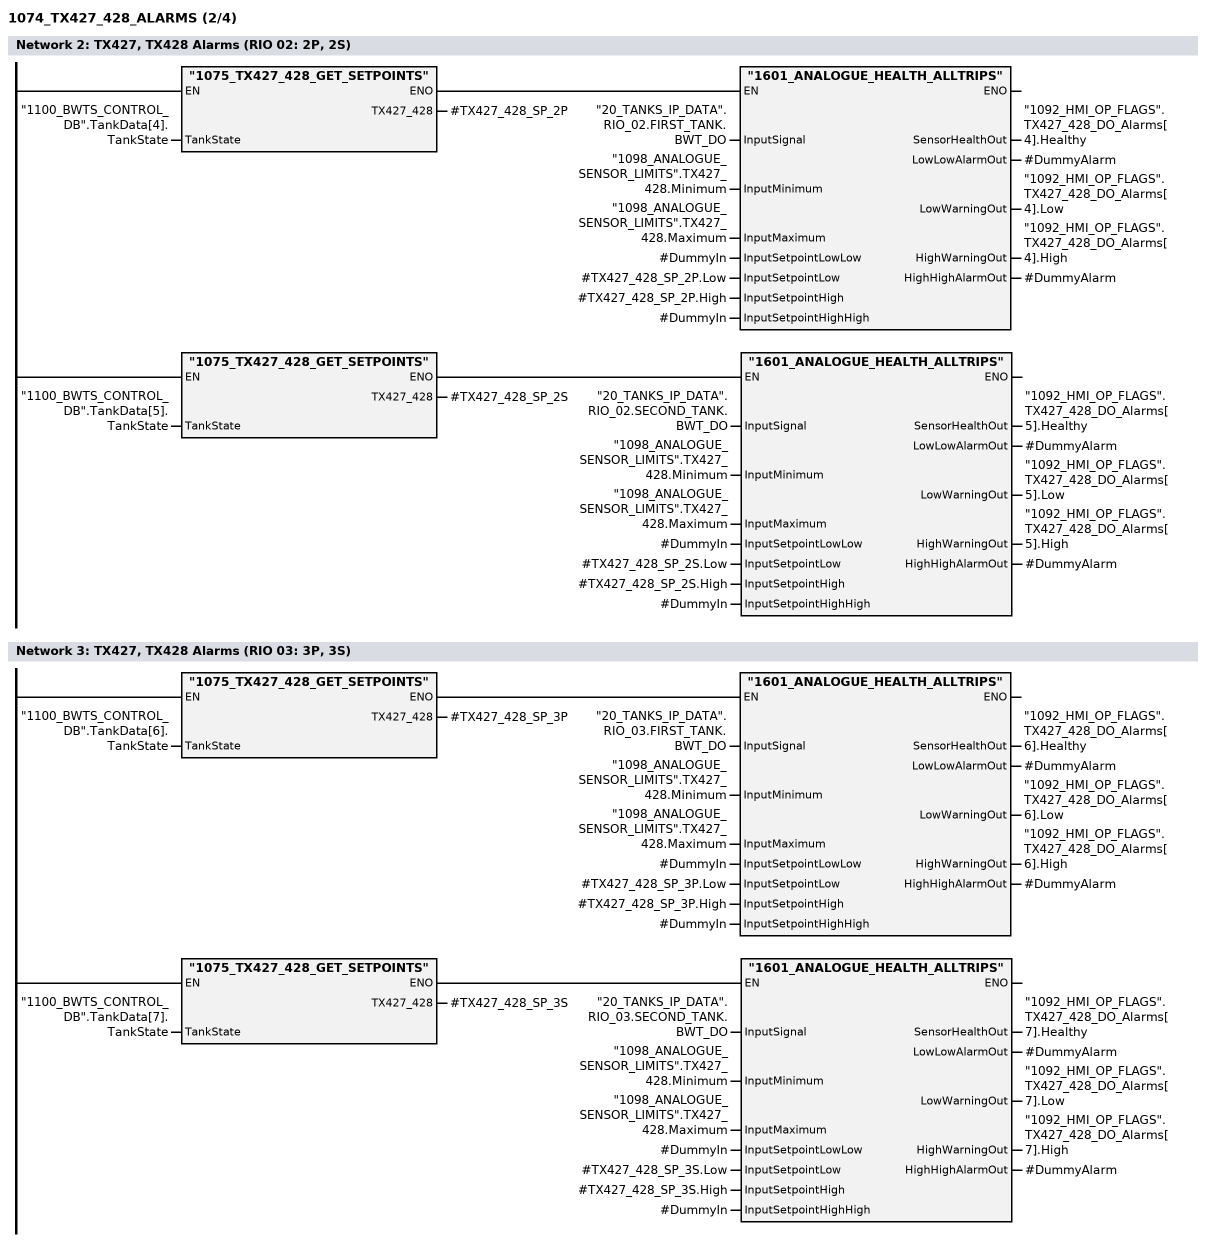
   RUNG wire#powerrail
      "1075_TX427_428_GET_SETPOINTS"(TankState := "1100_BWTS_CONTROL_DB".TankData[4].TankState, TX427_428 => #TX427_428_SP_2P)
      "1601_ANALOGUE_HEALTH_ALLTRIPS"(InputSignal := "20_TANKS_IP_DATA".RIO_02.FIRST_TANK.BWT_DO, InputMinimum := "1098_ANALOGUE_SENSOR_LIMITS".TX427_428.Minimum, InputMaximum := "1098_ANALOGUE_SENSOR_LIMITS".TX427_428.Maximum, InputSetpointLowLow := #DummyIn, InputSetpointLow := #TX427_428_SP_2P.Low, InputSetpointHigh := #TX427_428_SP_2P.High, InputSetpointHighHigh := #DummyIn, SensorHealthOut => "1092_HMI_OP_FLAGS".TX427_428_DO_Alarms[4].Healthy, LowLowAlarmOut => #DummyAlarm, LowWarningOut => "1092_HMI_OP_FLAGS".TX427_428_DO_Alarms[4].Low, HighWarningOut => "1092_HMI_OP_FLAGS".TX427_428_DO_Alarms[4].High, HighHighAlarmOut => #DummyAlarm)
   END_RUNG
   RUNG wire#powerrail
      "1075_TX427_428_GET_SETPOINTS"(TankState := "1100_BWTS_CONTROL_DB".TankData[5].TankState, TX427_428 => #TX427_428_SP_2S)
      "1601_ANALOGUE_HEALTH_ALLTRIPS"(InputSignal := "20_TANKS_IP_DATA".RIO_02.SECOND_TANK.BWT_DO, InputMinimum := "1098_ANALOGUE_SENSOR_LIMITS".TX427_428.Minimum, InputMaximum := "1098_ANALOGUE_SENSOR_LIMITS".TX427_428.Maximum, InputSetpointLowLow := #DummyIn, InputSetpointLow := #TX427_428_SP_2S.Low, InputSetpointHigh := #TX427_428_SP_2S.High, InputSetpointHighHigh := #DummyIn, SensorHealthOut => "1092_HMI_OP_FLAGS".TX427_428_DO_Alarms[5].Healthy, LowLowAlarmOut => #DummyAlarm, LowWarningOut => "1092_HMI_OP_FLAGS".TX427_428_DO_Alarms[5].Low, HighWarningOut => "1092_HMI_OP_FLAGS".TX427_428_DO_Alarms[5].High, HighHighAlarmOut => #DummyAlarm)
   END_RUNG
   // the same network as SCL:
   "1075_TX427_428_GET_SETPOINTS"(TankState := "1100_BWTS_CONTROL_DB".TankData[4].TankState,
                           TX427_428 => #TX427_428_SP_2P,
                           ENO => #_w1);
   IF #_w1 THEN
       "1601_ANALOGUE_HEALTH_ALLTRIPS"(InputSignal := "20_TANKS_IP_DATA".RIO_02.FIRST_TANK.BWT_DO,
                               InputMinimum := "1098_ANALOGUE_SENSOR_LIMITS".TX427_428.Minimum,
                               InputMaximum := "1098_ANALOGUE_SENSOR_LIMITS".TX427_428.Maximum,
                               InputSetpointLowLow := #DummyIn,
                               InputSetpointLow := #TX427_428_SP_2P.Low,
                               InputSetpointHigh := #TX427_428_SP_2P.High,
                               InputSetpointHighHigh := #DummyIn,
                               SensorHealthOut => "1092_HMI_OP_FLAGS".TX427_428_DO_Alarms[4].Healthy,
                               LowLowAlarmOut => #DummyAlarm,
                               LowWarningOut => "1092_HMI_OP_FLAGS".TX427_428_DO_Alarms[4].Low,
                               HighWarningOut => "1092_HMI_OP_FLAGS".TX427_428_DO_Alarms[4].High,
                               HighHighAlarmOut => #DummyAlarm);
   END_IF;
   "1075_TX427_428_GET_SETPOINTS"(TankState := "1100_BWTS_CONTROL_DB".TankData[5].TankState,
                           TX427_428 => #TX427_428_SP_2S,
                           ENO => #_w2);
   IF #_w2 THEN
       "1601_ANALOGUE_HEALTH_ALLTRIPS"(InputSignal := "20_TANKS_IP_DATA".RIO_02.SECOND_TANK.BWT_DO,
                               InputMinimum := "1098_ANALOGUE_SENSOR_LIMITS".TX427_428.Minimum,
                               InputMaximum := "1098_ANALOGUE_SENSOR_LIMITS".TX427_428.Maximum,
                               InputSetpointLowLow := #DummyIn,
                               InputSetpointLow := #TX427_428_SP_2S.Low,
                               InputSetpointHigh := #TX427_428_SP_2S.High,
                               InputSetpointHighHigh := #DummyIn,
                               SensorHealthOut => "1092_HMI_OP_FLAGS".TX427_428_DO_Alarms[5].Healthy,
                               LowLowAlarmOut => #DummyAlarm,
                               LowWarningOut => "1092_HMI_OP_FLAGS".TX427_428_DO_Alarms[5].Low,
                               HighWarningOut => "1092_HMI_OP_FLAGS".TX427_428_DO_Alarms[5].High,
                               HighHighAlarmOut => #DummyAlarm);
   END_IF;
END_REGION

REGION Network 3: TX427, TX428 Alarms (RIO 03: 3P, 3S)
   RUNG wire#powerrail
      "1075_TX427_428_GET_SETPOINTS"(TankState := "1100_BWTS_CONTROL_DB".TankData[6].TankState, TX427_428 => #TX427_428_SP_3P)
      "1601_ANALOGUE_HEALTH_ALLTRIPS"(InputSignal := "20_TANKS_IP_DATA".RIO_03.FIRST_TANK.BWT_DO, InputMinimum := "1098_ANALOGUE_SENSOR_LIMITS".TX427_428.Minimum, InputMaximum := "1098_ANALOGUE_SENSOR_LIMITS".TX427_428.Maximum, InputSetpointLowLow := #DummyIn, InputSetpointLow := #TX427_428_SP_3P.Low, InputSetpointHigh := #TX427_428_SP_3P.High, InputSetpointHighHigh := #DummyIn, SensorHealthOut => "1092_HMI_OP_FLAGS".TX427_428_DO_Alarms[6].Healthy, LowLowAlarmOut => #DummyAlarm, LowWarningOut => "1092_HMI_OP_FLAGS".TX427_428_DO_Alarms[6].Low, HighWarningOut => "1092_HMI_OP_FLAGS".TX427_428_DO_Alarms[6].High, HighHighAlarmOut => #DummyAlarm)
   END_RUNG
   RUNG wire#powerrail
      "1075_TX427_428_GET_SETPOINTS"(TankState := "1100_BWTS_CONTROL_DB".TankData[7].TankState, TX427_428 => #TX427_428_SP_3S)
      "1601_ANALOGUE_HEALTH_ALLTRIPS"(InputSignal := "20_TANKS_IP_DATA".RIO_03.SECOND_TANK.BWT_DO, InputMinimum := "1098_ANALOGUE_SENSOR_LIMITS".TX427_428.Minimum, InputMaximum := "1098_ANALOGUE_SENSOR_LIMITS".TX427_428.Maximum, InputSetpointLowLow := #DummyIn, InputSetpointLow := #TX427_428_SP_3S.Low, InputSetpointHigh := #TX427_428_SP_3S.High, InputSetpointHighHigh := #DummyIn, SensorHealthOut => "1092_HMI_OP_FLAGS".TX427_428_DO_Alarms[7].Healthy, LowLowAlarmOut => #DummyAlarm, LowWarningOut => "1092_HMI_OP_FLAGS".TX427_428_DO_Alarms[7].Low, HighWarningOut => "1092_HMI_OP_FLAGS".TX427_428_DO_Alarms[7].High, HighHighAlarmOut => #DummyAlarm)
   END_RUNG
   // the same network as SCL:
   "1075_TX427_428_GET_SETPOINTS"(TankState := "1100_BWTS_CONTROL_DB".TankData[6].TankState,
                           TX427_428 => #TX427_428_SP_3P,
                           ENO => #_w1);
   IF #_w1 THEN
       "1601_ANALOGUE_HEALTH_ALLTRIPS"(InputSignal := "20_TANKS_IP_DATA".RIO_03.FIRST_TANK.BWT_DO,
                               InputMinimum := "1098_ANALOGUE_SENSOR_LIMITS".TX427_428.Minimum,
                               InputMaximum := "1098_ANALOGUE_SENSOR_LIMITS".TX427_428.Maximum,
                               InputSetpointLowLow := #DummyIn,
                               InputSetpointLow := #TX427_428_SP_3P.Low,
                               InputSetpointHigh := #TX427_428_SP_3P.High,
                               InputSetpointHighHigh := #DummyIn,
                               SensorHealthOut => "1092_HMI_OP_FLAGS".TX427_428_DO_Alarms[6].Healthy,
                               LowLowAlarmOut => #DummyAlarm,
                               LowWarningOut => "1092_HMI_OP_FLAGS".TX427_428_DO_Alarms[6].Low,
                               HighWarningOut => "1092_HMI_OP_FLAGS".TX427_428_DO_Alarms[6].High,
                               HighHighAlarmOut => #DummyAlarm);
   END_IF;
   "1075_TX427_428_GET_SETPOINTS"(TankState := "1100_BWTS_CONTROL_DB".TankData[7].TankState,
                           TX427_428 => #TX427_428_SP_3S,
                           ENO => #_w2);
   IF #_w2 THEN
       "1601_ANALOGUE_HEALTH_ALLTRIPS"(InputSignal := "20_TANKS_IP_DATA".RIO_03.SECOND_TANK.BWT_DO,
                               InputMinimum := "1098_ANALOGUE_SENSOR_LIMITS".TX427_428.Minimum,
                               InputMaximum := "1098_ANALOGUE_SENSOR_LIMITS".TX427_428.Maximum,
                               InputSetpointLowLow := #DummyIn,
                               InputSetpointLow := #TX427_428_SP_3S.Low,
                               InputSetpointHigh := #TX427_428_SP_3S.High,
                               InputSetpointHighHigh := #DummyIn,
                               SensorHealthOut => "1092_HMI_OP_FLAGS".TX427_428_DO_Alarms[7].Healthy,
                               LowLowAlarmOut => #DummyAlarm,
                               LowWarningOut => "1092_HMI_OP_FLAGS".TX427_428_DO_Alarms[7].Low,
                               HighWarningOut => "1092_HMI_OP_FLAGS".TX427_428_DO_Alarms[7].High,
                               HighHighAlarmOut => #DummyAlarm);
   END_IF;
END_REGION

REGION Network 4: TX427, TX428 Alarms (RIO 04: 4P, 4S)
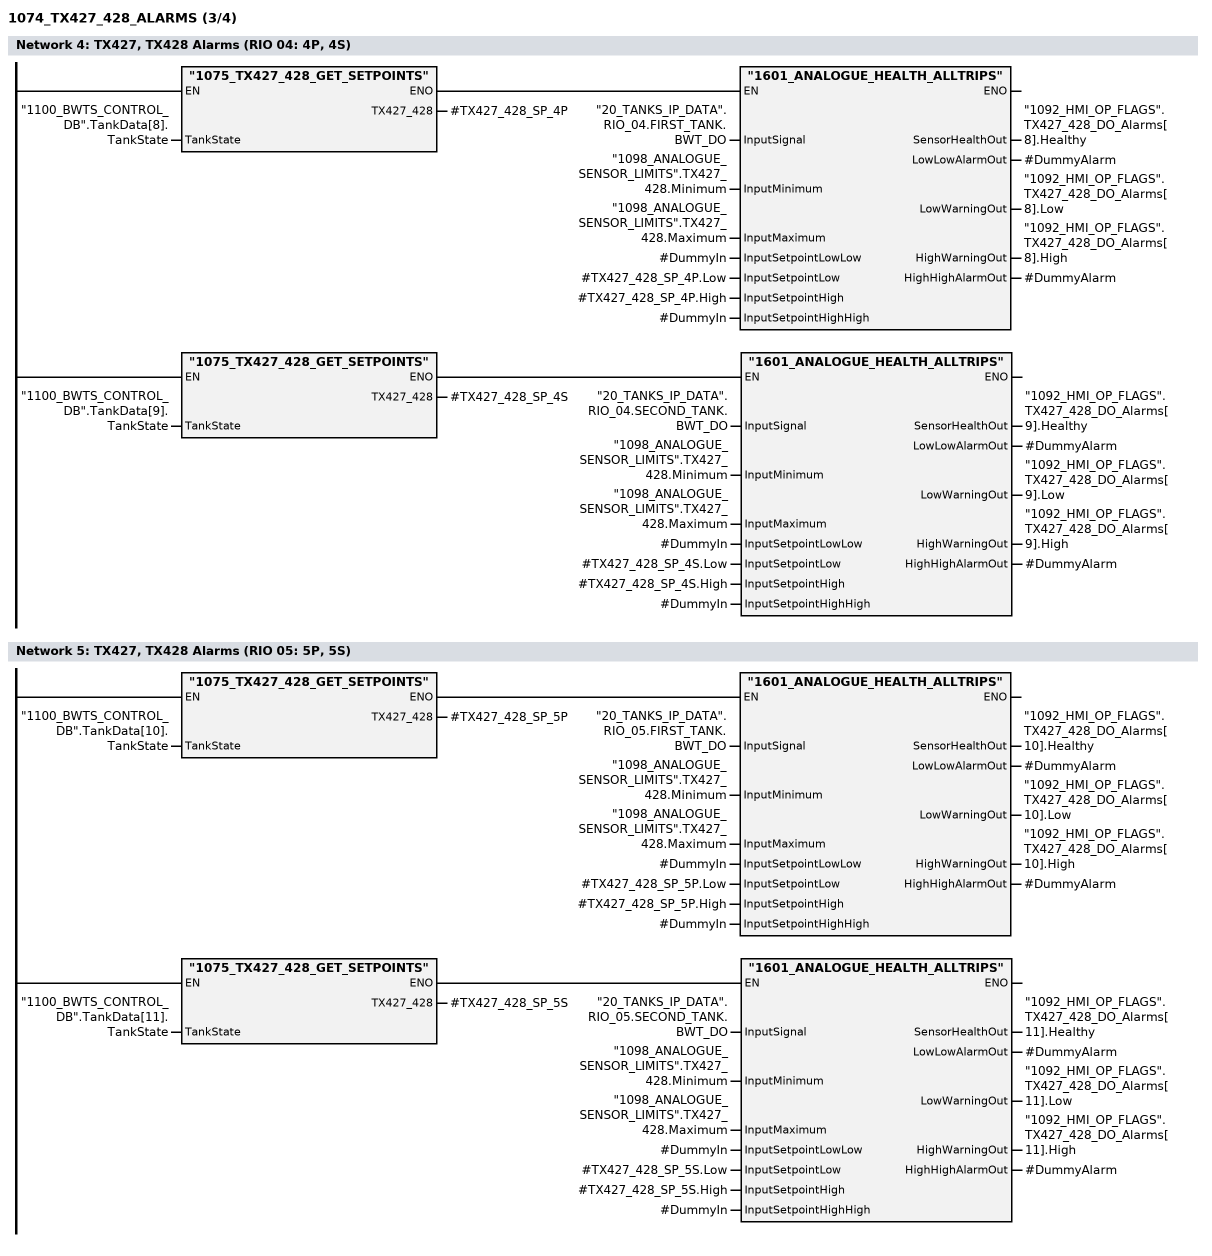
   RUNG wire#powerrail
      "1075_TX427_428_GET_SETPOINTS"(TankState := "1100_BWTS_CONTROL_DB".TankData[8].TankState, TX427_428 => #TX427_428_SP_4P)
      "1601_ANALOGUE_HEALTH_ALLTRIPS"(InputSignal := "20_TANKS_IP_DATA".RIO_04.FIRST_TANK.BWT_DO, InputMinimum := "1098_ANALOGUE_SENSOR_LIMITS".TX427_428.Minimum, InputMaximum := "1098_ANALOGUE_SENSOR_LIMITS".TX427_428.Maximum, InputSetpointLowLow := #DummyIn, InputSetpointLow := #TX427_428_SP_4P.Low, InputSetpointHigh := #TX427_428_SP_4P.High, InputSetpointHighHigh := #DummyIn, SensorHealthOut => "1092_HMI_OP_FLAGS".TX427_428_DO_Alarms[8].Healthy, LowLowAlarmOut => #DummyAlarm, LowWarningOut => "1092_HMI_OP_FLAGS".TX427_428_DO_Alarms[8].Low, HighWarningOut => "1092_HMI_OP_FLAGS".TX427_428_DO_Alarms[8].High, HighHighAlarmOut => #DummyAlarm)
   END_RUNG
   RUNG wire#powerrail
      "1075_TX427_428_GET_SETPOINTS"(TankState := "1100_BWTS_CONTROL_DB".TankData[9].TankState, TX427_428 => #TX427_428_SP_4S)
      "1601_ANALOGUE_HEALTH_ALLTRIPS"(InputSignal := "20_TANKS_IP_DATA".RIO_04.SECOND_TANK.BWT_DO, InputMinimum := "1098_ANALOGUE_SENSOR_LIMITS".TX427_428.Minimum, InputMaximum := "1098_ANALOGUE_SENSOR_LIMITS".TX427_428.Maximum, InputSetpointLowLow := #DummyIn, InputSetpointLow := #TX427_428_SP_4S.Low, InputSetpointHigh := #TX427_428_SP_4S.High, InputSetpointHighHigh := #DummyIn, SensorHealthOut => "1092_HMI_OP_FLAGS".TX427_428_DO_Alarms[9].Healthy, LowLowAlarmOut => #DummyAlarm, LowWarningOut => "1092_HMI_OP_FLAGS".TX427_428_DO_Alarms[9].Low, HighWarningOut => "1092_HMI_OP_FLAGS".TX427_428_DO_Alarms[9].High, HighHighAlarmOut => #DummyAlarm)
   END_RUNG
   // the same network as SCL:
   "1075_TX427_428_GET_SETPOINTS"(TankState := "1100_BWTS_CONTROL_DB".TankData[8].TankState,
                           TX427_428 => #TX427_428_SP_4P,
                           ENO => #_w1);
   IF #_w1 THEN
       "1601_ANALOGUE_HEALTH_ALLTRIPS"(InputSignal := "20_TANKS_IP_DATA".RIO_04.FIRST_TANK.BWT_DO,
                               InputMinimum := "1098_ANALOGUE_SENSOR_LIMITS".TX427_428.Minimum,
                               InputMaximum := "1098_ANALOGUE_SENSOR_LIMITS".TX427_428.Maximum,
                               InputSetpointLowLow := #DummyIn,
                               InputSetpointLow := #TX427_428_SP_4P.Low,
                               InputSetpointHigh := #TX427_428_SP_4P.High,
                               InputSetpointHighHigh := #DummyIn,
                               SensorHealthOut => "1092_HMI_OP_FLAGS".TX427_428_DO_Alarms[8].Healthy,
                               LowLowAlarmOut => #DummyAlarm,
                               LowWarningOut => "1092_HMI_OP_FLAGS".TX427_428_DO_Alarms[8].Low,
                               HighWarningOut => "1092_HMI_OP_FLAGS".TX427_428_DO_Alarms[8].High,
                               HighHighAlarmOut => #DummyAlarm);
   END_IF;
   "1075_TX427_428_GET_SETPOINTS"(TankState := "1100_BWTS_CONTROL_DB".TankData[9].TankState,
                           TX427_428 => #TX427_428_SP_4S,
                           ENO => #_w2);
   IF #_w2 THEN
       "1601_ANALOGUE_HEALTH_ALLTRIPS"(InputSignal := "20_TANKS_IP_DATA".RIO_04.SECOND_TANK.BWT_DO,
                               InputMinimum := "1098_ANALOGUE_SENSOR_LIMITS".TX427_428.Minimum,
                               InputMaximum := "1098_ANALOGUE_SENSOR_LIMITS".TX427_428.Maximum,
                               InputSetpointLowLow := #DummyIn,
                               InputSetpointLow := #TX427_428_SP_4S.Low,
                               InputSetpointHigh := #TX427_428_SP_4S.High,
                               InputSetpointHighHigh := #DummyIn,
                               SensorHealthOut => "1092_HMI_OP_FLAGS".TX427_428_DO_Alarms[9].Healthy,
                               LowLowAlarmOut => #DummyAlarm,
                               LowWarningOut => "1092_HMI_OP_FLAGS".TX427_428_DO_Alarms[9].Low,
                               HighWarningOut => "1092_HMI_OP_FLAGS".TX427_428_DO_Alarms[9].High,
                               HighHighAlarmOut => #DummyAlarm);
   END_IF;
END_REGION

REGION Network 5: TX427, TX428 Alarms (RIO 05: 5P, 5S)
   RUNG wire#powerrail
      "1075_TX427_428_GET_SETPOINTS"(TankState := "1100_BWTS_CONTROL_DB".TankData[10].TankState, TX427_428 => #TX427_428_SP_5P)
      "1601_ANALOGUE_HEALTH_ALLTRIPS"(InputSignal := "20_TANKS_IP_DATA".RIO_05.FIRST_TANK.BWT_DO, InputMinimum := "1098_ANALOGUE_SENSOR_LIMITS".TX427_428.Minimum, InputMaximum := "1098_ANALOGUE_SENSOR_LIMITS".TX427_428.Maximum, InputSetpointLowLow := #DummyIn, InputSetpointLow := #TX427_428_SP_5P.Low, InputSetpointHigh := #TX427_428_SP_5P.High, InputSetpointHighHigh := #DummyIn, SensorHealthOut => "1092_HMI_OP_FLAGS".TX427_428_DO_Alarms[10].Healthy, LowLowAlarmOut => #DummyAlarm, LowWarningOut => "1092_HMI_OP_FLAGS".TX427_428_DO_Alarms[10].Low, HighWarningOut => "1092_HMI_OP_FLAGS".TX427_428_DO_Alarms[10].High, HighHighAlarmOut => #DummyAlarm)
   END_RUNG
   RUNG wire#powerrail
      "1075_TX427_428_GET_SETPOINTS"(TankState := "1100_BWTS_CONTROL_DB".TankData[11].TankState, TX427_428 => #TX427_428_SP_5S)
      "1601_ANALOGUE_HEALTH_ALLTRIPS"(InputSignal := "20_TANKS_IP_DATA".RIO_05.SECOND_TANK.BWT_DO, InputMinimum := "1098_ANALOGUE_SENSOR_LIMITS".TX427_428.Minimum, InputMaximum := "1098_ANALOGUE_SENSOR_LIMITS".TX427_428.Maximum, InputSetpointLowLow := #DummyIn, InputSetpointLow := #TX427_428_SP_5S.Low, InputSetpointHigh := #TX427_428_SP_5S.High, InputSetpointHighHigh := #DummyIn, SensorHealthOut => "1092_HMI_OP_FLAGS".TX427_428_DO_Alarms[11].Healthy, LowLowAlarmOut => #DummyAlarm, LowWarningOut => "1092_HMI_OP_FLAGS".TX427_428_DO_Alarms[11].Low, HighWarningOut => "1092_HMI_OP_FLAGS".TX427_428_DO_Alarms[11].High, HighHighAlarmOut => #DummyAlarm)
   END_RUNG
   // the same network as SCL:
   "1075_TX427_428_GET_SETPOINTS"(TankState := "1100_BWTS_CONTROL_DB".TankData[10].TankState,
                           TX427_428 => #TX427_428_SP_5P,
                           ENO => #_w1);
   IF #_w1 THEN
       "1601_ANALOGUE_HEALTH_ALLTRIPS"(InputSignal := "20_TANKS_IP_DATA".RIO_05.FIRST_TANK.BWT_DO,
                               InputMinimum := "1098_ANALOGUE_SENSOR_LIMITS".TX427_428.Minimum,
                               InputMaximum := "1098_ANALOGUE_SENSOR_LIMITS".TX427_428.Maximum,
                               InputSetpointLowLow := #DummyIn,
                               InputSetpointLow := #TX427_428_SP_5P.Low,
                               InputSetpointHigh := #TX427_428_SP_5P.High,
                               InputSetpointHighHigh := #DummyIn,
                               SensorHealthOut => "1092_HMI_OP_FLAGS".TX427_428_DO_Alarms[10].Healthy,
                               LowLowAlarmOut => #DummyAlarm,
                               LowWarningOut => "1092_HMI_OP_FLAGS".TX427_428_DO_Alarms[10].Low,
                               HighWarningOut => "1092_HMI_OP_FLAGS".TX427_428_DO_Alarms[10].High,
                               HighHighAlarmOut => #DummyAlarm);
   END_IF;
   "1075_TX427_428_GET_SETPOINTS"(TankState := "1100_BWTS_CONTROL_DB".TankData[11].TankState,
                           TX427_428 => #TX427_428_SP_5S,
                           ENO => #_w2);
   IF #_w2 THEN
       "1601_ANALOGUE_HEALTH_ALLTRIPS"(InputSignal := "20_TANKS_IP_DATA".RIO_05.SECOND_TANK.BWT_DO,
                               InputMinimum := "1098_ANALOGUE_SENSOR_LIMITS".TX427_428.Minimum,
                               InputMaximum := "1098_ANALOGUE_SENSOR_LIMITS".TX427_428.Maximum,
                               InputSetpointLowLow := #DummyIn,
                               InputSetpointLow := #TX427_428_SP_5S.Low,
                               InputSetpointHigh := #TX427_428_SP_5S.High,
                               InputSetpointHighHigh := #DummyIn,
                               SensorHealthOut => "1092_HMI_OP_FLAGS".TX427_428_DO_Alarms[11].Healthy,
                               LowLowAlarmOut => #DummyAlarm,
                               LowWarningOut => "1092_HMI_OP_FLAGS".TX427_428_DO_Alarms[11].Low,
                               HighWarningOut => "1092_HMI_OP_FLAGS".TX427_428_DO_Alarms[11].High,
                               HighHighAlarmOut => #DummyAlarm);
   END_IF;
END_REGION

REGION Network 6: TX427, TX428 Alarms (RIO 06: 6P, 6S)
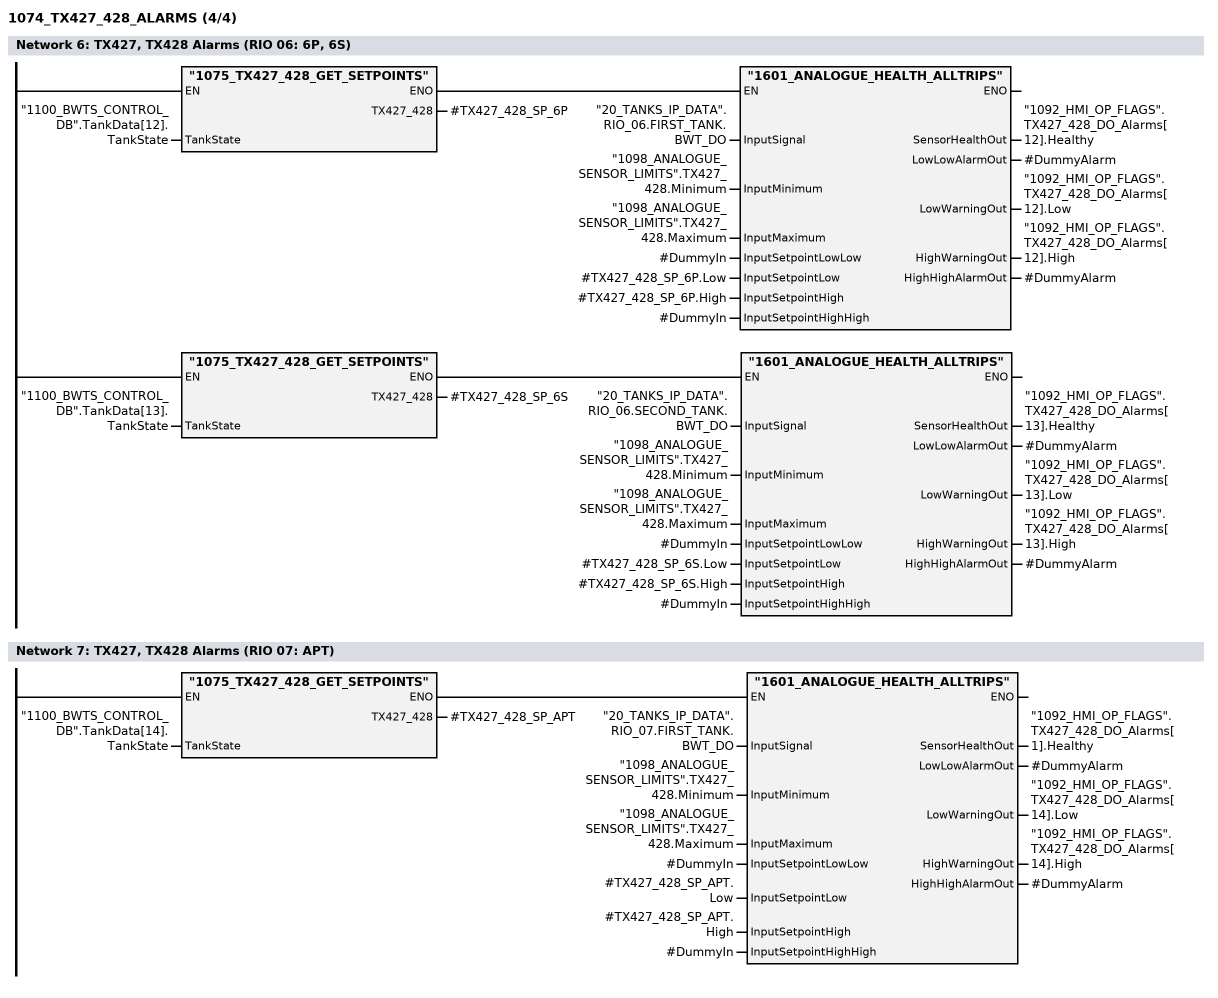
   RUNG wire#powerrail
      "1075_TX427_428_GET_SETPOINTS"(TankState := "1100_BWTS_CONTROL_DB".TankData[12].TankState, TX427_428 => #TX427_428_SP_6P)
      "1601_ANALOGUE_HEALTH_ALLTRIPS"(InputSignal := "20_TANKS_IP_DATA".RIO_06.FIRST_TANK.BWT_DO, InputMinimum := "1098_ANALOGUE_SENSOR_LIMITS".TX427_428.Minimum, InputMaximum := "1098_ANALOGUE_SENSOR_LIMITS".TX427_428.Maximum, InputSetpointLowLow := #DummyIn, InputSetpointLow := #TX427_428_SP_6P.Low, InputSetpointHigh := #TX427_428_SP_6P.High, InputSetpointHighHigh := #DummyIn, SensorHealthOut => "1092_HMI_OP_FLAGS".TX427_428_DO_Alarms[12].Healthy, LowLowAlarmOut => #DummyAlarm, LowWarningOut => "1092_HMI_OP_FLAGS".TX427_428_DO_Alarms[12].Low, HighWarningOut => "1092_HMI_OP_FLAGS".TX427_428_DO_Alarms[12].High, HighHighAlarmOut => #DummyAlarm)
   END_RUNG
   RUNG wire#powerrail
      "1075_TX427_428_GET_SETPOINTS"(TankState := "1100_BWTS_CONTROL_DB".TankData[13].TankState, TX427_428 => #TX427_428_SP_6S)
      "1601_ANALOGUE_HEALTH_ALLTRIPS"(InputSignal := "20_TANKS_IP_DATA".RIO_06.SECOND_TANK.BWT_DO, InputMinimum := "1098_ANALOGUE_SENSOR_LIMITS".TX427_428.Minimum, InputMaximum := "1098_ANALOGUE_SENSOR_LIMITS".TX427_428.Maximum, InputSetpointLowLow := #DummyIn, InputSetpointLow := #TX427_428_SP_6S.Low, InputSetpointHigh := #TX427_428_SP_6S.High, InputSetpointHighHigh := #DummyIn, SensorHealthOut => "1092_HMI_OP_FLAGS".TX427_428_DO_Alarms[13].Healthy, LowLowAlarmOut => #DummyAlarm, LowWarningOut => "1092_HMI_OP_FLAGS".TX427_428_DO_Alarms[13].Low, HighWarningOut => "1092_HMI_OP_FLAGS".TX427_428_DO_Alarms[13].High, HighHighAlarmOut => #DummyAlarm)
   END_RUNG
   // the same network as SCL:
   "1075_TX427_428_GET_SETPOINTS"(TankState := "1100_BWTS_CONTROL_DB".TankData[12].TankState,
                           TX427_428 => #TX427_428_SP_6P,
                           ENO => #_w1);
   IF #_w1 THEN
       "1601_ANALOGUE_HEALTH_ALLTRIPS"(InputSignal := "20_TANKS_IP_DATA".RIO_06.FIRST_TANK.BWT_DO,
                               InputMinimum := "1098_ANALOGUE_SENSOR_LIMITS".TX427_428.Minimum,
                               InputMaximum := "1098_ANALOGUE_SENSOR_LIMITS".TX427_428.Maximum,
                               InputSetpointLowLow := #DummyIn,
                               InputSetpointLow := #TX427_428_SP_6P.Low,
                               InputSetpointHigh := #TX427_428_SP_6P.High,
                               InputSetpointHighHigh := #DummyIn,
                               SensorHealthOut => "1092_HMI_OP_FLAGS".TX427_428_DO_Alarms[12].Healthy,
                               LowLowAlarmOut => #DummyAlarm,
                               LowWarningOut => "1092_HMI_OP_FLAGS".TX427_428_DO_Alarms[12].Low,
                               HighWarningOut => "1092_HMI_OP_FLAGS".TX427_428_DO_Alarms[12].High,
                               HighHighAlarmOut => #DummyAlarm);
   END_IF;
   "1075_TX427_428_GET_SETPOINTS"(TankState := "1100_BWTS_CONTROL_DB".TankData[13].TankState,
                           TX427_428 => #TX427_428_SP_6S,
                           ENO => #_w2);
   IF #_w2 THEN
       "1601_ANALOGUE_HEALTH_ALLTRIPS"(InputSignal := "20_TANKS_IP_DATA".RIO_06.SECOND_TANK.BWT_DO,
                               InputMinimum := "1098_ANALOGUE_SENSOR_LIMITS".TX427_428.Minimum,
                               InputMaximum := "1098_ANALOGUE_SENSOR_LIMITS".TX427_428.Maximum,
                               InputSetpointLowLow := #DummyIn,
                               InputSetpointLow := #TX427_428_SP_6S.Low,
                               InputSetpointHigh := #TX427_428_SP_6S.High,
                               InputSetpointHighHigh := #DummyIn,
                               SensorHealthOut => "1092_HMI_OP_FLAGS".TX427_428_DO_Alarms[13].Healthy,
                               LowLowAlarmOut => #DummyAlarm,
                               LowWarningOut => "1092_HMI_OP_FLAGS".TX427_428_DO_Alarms[13].Low,
                               HighWarningOut => "1092_HMI_OP_FLAGS".TX427_428_DO_Alarms[13].High,
                               HighHighAlarmOut => #DummyAlarm);
   END_IF;
END_REGION

REGION Network 7: TX427, TX428 Alarms (RIO 07: APT)
   RUNG wire#powerrail
      "1075_TX427_428_GET_SETPOINTS"(TankState := "1100_BWTS_CONTROL_DB".TankData[14].TankState, TX427_428 => #TX427_428_SP_APT)
      "1601_ANALOGUE_HEALTH_ALLTRIPS"(InputSignal := "20_TANKS_IP_DATA".RIO_07.FIRST_TANK.BWT_DO, InputMinimum := "1098_ANALOGUE_SENSOR_LIMITS".TX427_428.Minimum, InputMaximum := "1098_ANALOGUE_SENSOR_LIMITS".TX427_428.Maximum, InputSetpointLowLow := #DummyIn, InputSetpointLow := #TX427_428_SP_APT.Low, InputSetpointHigh := #TX427_428_SP_APT.High, InputSetpointHighHigh := #DummyIn, SensorHealthOut => "1092_HMI_OP_FLAGS".TX427_428_DO_Alarms[1].Healthy, LowLowAlarmOut => #DummyAlarm, LowWarningOut => "1092_HMI_OP_FLAGS".TX427_428_DO_Alarms[14].Low, HighWarningOut => "1092_HMI_OP_FLAGS".TX427_428_DO_Alarms[14].High, HighHighAlarmOut => #DummyAlarm)
   END_RUNG
   // the same network as SCL:
   "1075_TX427_428_GET_SETPOINTS"(TankState := "1100_BWTS_CONTROL_DB".TankData[14].TankState,
                           TX427_428 => #TX427_428_SP_APT,
                           ENO => #_w1);
   IF #_w1 THEN
       "1601_ANALOGUE_HEALTH_ALLTRIPS"(InputSignal := "20_TANKS_IP_DATA".RIO_07.FIRST_TANK.BWT_DO,
                               InputMinimum := "1098_ANALOGUE_SENSOR_LIMITS".TX427_428.Minimum,
                               InputMaximum := "1098_ANALOGUE_SENSOR_LIMITS".TX427_428.Maximum,
                               InputSetpointLowLow := #DummyIn,
                               InputSetpointLow := #TX427_428_SP_APT.Low,
                               InputSetpointHigh := #TX427_428_SP_APT.High,
                               InputSetpointHighHigh := #DummyIn,
                               SensorHealthOut => "1092_HMI_OP_FLAGS".TX427_428_DO_Alarms[1].Healthy,
                               LowLowAlarmOut => #DummyAlarm,
                               LowWarningOut => "1092_HMI_OP_FLAGS".TX427_428_DO_Alarms[14].Low,
                               HighWarningOut => "1092_HMI_OP_FLAGS".TX427_428_DO_Alarms[14].High,
                               HighHighAlarmOut => #DummyAlarm);
   END_IF;
END_REGION
END_FUNCTION

FUNCTION "1075_TX427_428_GET_SETPOINTS" : Void   // FC1075, SCL
{ S7_Optimized_Access := 'TRUE' }
VERSION : 0.1
   VAR_INPUT
      TankState : Int;
   END_VAR
   VAR_OUTPUT
      TX427_428 : "ANALOG_SENSOR_SETPOINTS";
   END_VAR
   VAR CONSTANT
      TankState_Init : Int := 1000;
      TankState_PreDwell : Int := 1001;
      TankState_DeOx : Int := 1002;
      TankState_MidDwell : Int := 1003;
      TankState_ReOx : Int := 1004;
      TankState_PostDwell : Int := 1005;
      TankState_Done : Int := 1006;
   END_VAR
BEGIN
   (* This function is required to define the setpoints of the DO sensors based on the current state.
       The alarms shall use differing setpoints in different phases defined as:
       DEOX alarm setpoints if in DeOx, or Mid-Dwell
       REOX alarm setpoints if in PreDwell, Reox, or PostDwell (All others values) *)

   IF #TankState = #TankState_DeOx OR #TankState = #TankState_MidDwell THEN
       #TX427_428 := "1094_ANALOGUE_SENSOR_SETPOINTS".TX427_428_DEOX;
   ELSE
       #TX427_428 := "1094_ANALOGUE_SENSOR_SETPOINTS".TX427_428_REOX;
   END_IF;
END_FUNCTION

FUNCTION "1076_LS425_442_ALARMS" : Void   // FC1076, LAD
{ S7_Optimized_Access := 'TRUE' }
VERSION : 0.1
// Alarm wrapper function for BWT Level Switch on each tank.
   VAR CONSTANT
      InputTripLevel : Bool;   // The input trip level for this function, if the input is equal to this digital value, trip the alarm.
   END_VAR
BEGIN

REGION Network 1: LS425, LS442 Alarms (RIO 01: FPT. 1P, 1S)
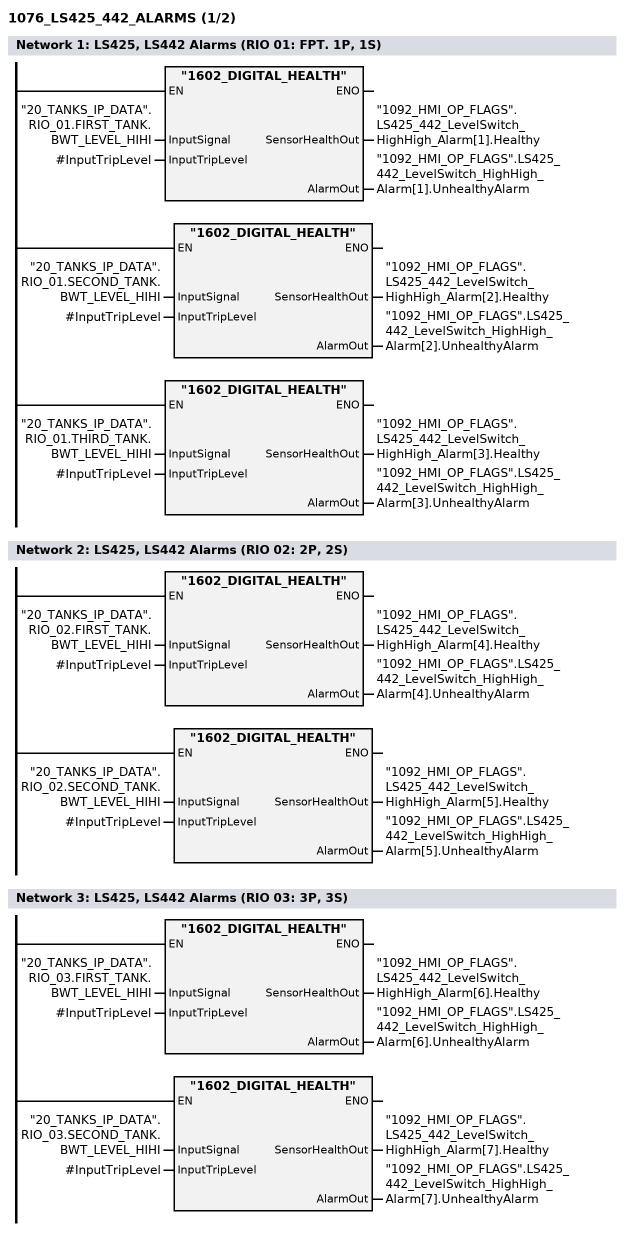
   RUNG wire#powerrail
      "1602_DIGITAL_HEALTH"(InputSignal := "20_TANKS_IP_DATA".RIO_01.FIRST_TANK.BWT_LEVEL_HIHI, InputTripLevel := #InputTripLevel, SensorHealthOut => "1092_HMI_OP_FLAGS".LS425_442_LevelSwitch_HighHigh_Alarm[1].Healthy, AlarmOut => "1092_HMI_OP_FLAGS".LS425_442_LevelSwitch_HighHigh_Alarm[1].UnhealthyAlarm)
   END_RUNG
   RUNG wire#powerrail
      "1602_DIGITAL_HEALTH"(InputSignal := "20_TANKS_IP_DATA".RIO_01.SECOND_TANK.BWT_LEVEL_HIHI, InputTripLevel := #InputTripLevel, SensorHealthOut => "1092_HMI_OP_FLAGS".LS425_442_LevelSwitch_HighHigh_Alarm[2].Healthy, AlarmOut => "1092_HMI_OP_FLAGS".LS425_442_LevelSwitch_HighHigh_Alarm[2].UnhealthyAlarm)
   END_RUNG
   RUNG wire#powerrail
      "1602_DIGITAL_HEALTH"(InputSignal := "20_TANKS_IP_DATA".RIO_01.THIRD_TANK.BWT_LEVEL_HIHI, InputTripLevel := #InputTripLevel, SensorHealthOut => "1092_HMI_OP_FLAGS".LS425_442_LevelSwitch_HighHigh_Alarm[3].Healthy, AlarmOut => "1092_HMI_OP_FLAGS".LS425_442_LevelSwitch_HighHigh_Alarm[3].UnhealthyAlarm)
   END_RUNG
   // the same network as SCL:
   "1602_DIGITAL_HEALTH"(InputSignal := "20_TANKS_IP_DATA".RIO_01.FIRST_TANK.BWT_LEVEL_HIHI,
                         InputTripLevel := #InputTripLevel,
                         SensorHealthOut => "1092_HMI_OP_FLAGS".LS425_442_LevelSwitch_HighHigh_Alarm[1].Healthy,
                         AlarmOut => "1092_HMI_OP_FLAGS".LS425_442_LevelSwitch_HighHigh_Alarm[1].UnhealthyAlarm);
   "1602_DIGITAL_HEALTH"(InputSignal := "20_TANKS_IP_DATA".RIO_01.SECOND_TANK.BWT_LEVEL_HIHI,
                         InputTripLevel := #InputTripLevel,
                         SensorHealthOut => "1092_HMI_OP_FLAGS".LS425_442_LevelSwitch_HighHigh_Alarm[2].Healthy,
                         AlarmOut => "1092_HMI_OP_FLAGS".LS425_442_LevelSwitch_HighHigh_Alarm[2].UnhealthyAlarm);
   "1602_DIGITAL_HEALTH"(InputSignal := "20_TANKS_IP_DATA".RIO_01.THIRD_TANK.BWT_LEVEL_HIHI,
                         InputTripLevel := #InputTripLevel,
                         SensorHealthOut => "1092_HMI_OP_FLAGS".LS425_442_LevelSwitch_HighHigh_Alarm[3].Healthy,
                         AlarmOut => "1092_HMI_OP_FLAGS".LS425_442_LevelSwitch_HighHigh_Alarm[3].UnhealthyAlarm);
END_REGION

REGION Network 2: LS425, LS442 Alarms (RIO 02: 2P, 2S)
   RUNG wire#powerrail
      "1602_DIGITAL_HEALTH"(InputSignal := "20_TANKS_IP_DATA".RIO_02.FIRST_TANK.BWT_LEVEL_HIHI, InputTripLevel := #InputTripLevel, SensorHealthOut => "1092_HMI_OP_FLAGS".LS425_442_LevelSwitch_HighHigh_Alarm[4].Healthy, AlarmOut => "1092_HMI_OP_FLAGS".LS425_442_LevelSwitch_HighHigh_Alarm[4].UnhealthyAlarm)
   END_RUNG
   RUNG wire#powerrail
      "1602_DIGITAL_HEALTH"(InputSignal := "20_TANKS_IP_DATA".RIO_02.SECOND_TANK.BWT_LEVEL_HIHI, InputTripLevel := #InputTripLevel, SensorHealthOut => "1092_HMI_OP_FLAGS".LS425_442_LevelSwitch_HighHigh_Alarm[5].Healthy, AlarmOut => "1092_HMI_OP_FLAGS".LS425_442_LevelSwitch_HighHigh_Alarm[5].UnhealthyAlarm)
   END_RUNG
   // the same network as SCL:
   "1602_DIGITAL_HEALTH"(InputSignal := "20_TANKS_IP_DATA".RIO_02.FIRST_TANK.BWT_LEVEL_HIHI,
                         InputTripLevel := #InputTripLevel,
                         SensorHealthOut => "1092_HMI_OP_FLAGS".LS425_442_LevelSwitch_HighHigh_Alarm[4].Healthy,
                         AlarmOut => "1092_HMI_OP_FLAGS".LS425_442_LevelSwitch_HighHigh_Alarm[4].UnhealthyAlarm);
   "1602_DIGITAL_HEALTH"(InputSignal := "20_TANKS_IP_DATA".RIO_02.SECOND_TANK.BWT_LEVEL_HIHI,
                         InputTripLevel := #InputTripLevel,
                         SensorHealthOut => "1092_HMI_OP_FLAGS".LS425_442_LevelSwitch_HighHigh_Alarm[5].Healthy,
                         AlarmOut => "1092_HMI_OP_FLAGS".LS425_442_LevelSwitch_HighHigh_Alarm[5].UnhealthyAlarm);
END_REGION

REGION Network 3: LS425, LS442 Alarms (RIO 03: 3P, 3S)
   RUNG wire#powerrail
      "1602_DIGITAL_HEALTH"(InputSignal := "20_TANKS_IP_DATA".RIO_03.FIRST_TANK.BWT_LEVEL_HIHI, InputTripLevel := #InputTripLevel, SensorHealthOut => "1092_HMI_OP_FLAGS".LS425_442_LevelSwitch_HighHigh_Alarm[6].Healthy, AlarmOut => "1092_HMI_OP_FLAGS".LS425_442_LevelSwitch_HighHigh_Alarm[6].UnhealthyAlarm)
   END_RUNG
   RUNG wire#powerrail
      "1602_DIGITAL_HEALTH"(InputSignal := "20_TANKS_IP_DATA".RIO_03.SECOND_TANK.BWT_LEVEL_HIHI, InputTripLevel := #InputTripLevel, SensorHealthOut => "1092_HMI_OP_FLAGS".LS425_442_LevelSwitch_HighHigh_Alarm[7].Healthy, AlarmOut => "1092_HMI_OP_FLAGS".LS425_442_LevelSwitch_HighHigh_Alarm[7].UnhealthyAlarm)
   END_RUNG
   // the same network as SCL:
   "1602_DIGITAL_HEALTH"(InputSignal := "20_TANKS_IP_DATA".RIO_03.FIRST_TANK.BWT_LEVEL_HIHI,
                         InputTripLevel := #InputTripLevel,
                         SensorHealthOut => "1092_HMI_OP_FLAGS".LS425_442_LevelSwitch_HighHigh_Alarm[6].Healthy,
                         AlarmOut => "1092_HMI_OP_FLAGS".LS425_442_LevelSwitch_HighHigh_Alarm[6].UnhealthyAlarm);
   "1602_DIGITAL_HEALTH"(InputSignal := "20_TANKS_IP_DATA".RIO_03.SECOND_TANK.BWT_LEVEL_HIHI,
                         InputTripLevel := #InputTripLevel,
                         SensorHealthOut => "1092_HMI_OP_FLAGS".LS425_442_LevelSwitch_HighHigh_Alarm[7].Healthy,
                         AlarmOut => "1092_HMI_OP_FLAGS".LS425_442_LevelSwitch_HighHigh_Alarm[7].UnhealthyAlarm);
END_REGION

REGION Network 4: LS425, LS442 Alarms (RIO 04: 4P, 4S)
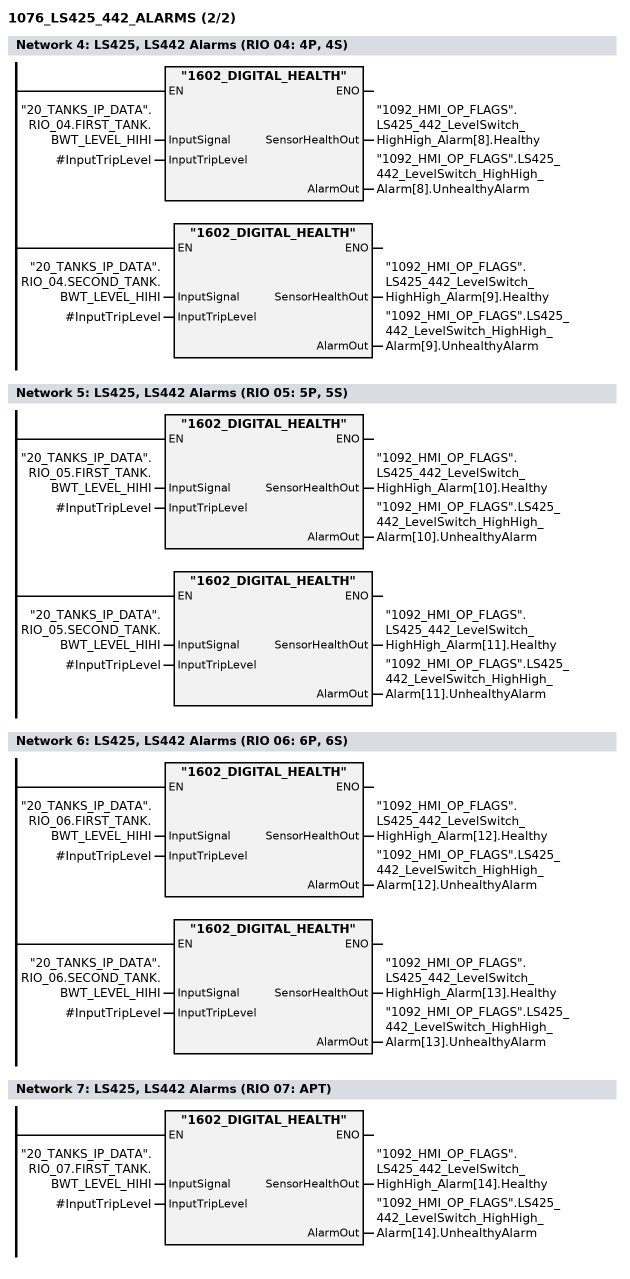
   RUNG wire#powerrail
      "1602_DIGITAL_HEALTH"(InputSignal := "20_TANKS_IP_DATA".RIO_04.FIRST_TANK.BWT_LEVEL_HIHI, InputTripLevel := #InputTripLevel, SensorHealthOut => "1092_HMI_OP_FLAGS".LS425_442_LevelSwitch_HighHigh_Alarm[8].Healthy, AlarmOut => "1092_HMI_OP_FLAGS".LS425_442_LevelSwitch_HighHigh_Alarm[8].UnhealthyAlarm)
   END_RUNG
   RUNG wire#powerrail
      "1602_DIGITAL_HEALTH"(InputSignal := "20_TANKS_IP_DATA".RIO_04.SECOND_TANK.BWT_LEVEL_HIHI, InputTripLevel := #InputTripLevel, SensorHealthOut => "1092_HMI_OP_FLAGS".LS425_442_LevelSwitch_HighHigh_Alarm[9].Healthy, AlarmOut => "1092_HMI_OP_FLAGS".LS425_442_LevelSwitch_HighHigh_Alarm[9].UnhealthyAlarm)
   END_RUNG
   // the same network as SCL:
   "1602_DIGITAL_HEALTH"(InputSignal := "20_TANKS_IP_DATA".RIO_04.FIRST_TANK.BWT_LEVEL_HIHI,
                         InputTripLevel := #InputTripLevel,
                         SensorHealthOut => "1092_HMI_OP_FLAGS".LS425_442_LevelSwitch_HighHigh_Alarm[8].Healthy,
                         AlarmOut => "1092_HMI_OP_FLAGS".LS425_442_LevelSwitch_HighHigh_Alarm[8].UnhealthyAlarm);
   "1602_DIGITAL_HEALTH"(InputSignal := "20_TANKS_IP_DATA".RIO_04.SECOND_TANK.BWT_LEVEL_HIHI,
                         InputTripLevel := #InputTripLevel,
                         SensorHealthOut => "1092_HMI_OP_FLAGS".LS425_442_LevelSwitch_HighHigh_Alarm[9].Healthy,
                         AlarmOut => "1092_HMI_OP_FLAGS".LS425_442_LevelSwitch_HighHigh_Alarm[9].UnhealthyAlarm);
END_REGION

REGION Network 5: LS425, LS442 Alarms (RIO 05: 5P, 5S)
   RUNG wire#powerrail
      "1602_DIGITAL_HEALTH"(InputSignal := "20_TANKS_IP_DATA".RIO_05.FIRST_TANK.BWT_LEVEL_HIHI, InputTripLevel := #InputTripLevel, SensorHealthOut => "1092_HMI_OP_FLAGS".LS425_442_LevelSwitch_HighHigh_Alarm[10].Healthy, AlarmOut => "1092_HMI_OP_FLAGS".LS425_442_LevelSwitch_HighHigh_Alarm[10].UnhealthyAlarm)
   END_RUNG
   RUNG wire#powerrail
      "1602_DIGITAL_HEALTH"(InputSignal := "20_TANKS_IP_DATA".RIO_05.SECOND_TANK.BWT_LEVEL_HIHI, InputTripLevel := #InputTripLevel, SensorHealthOut => "1092_HMI_OP_FLAGS".LS425_442_LevelSwitch_HighHigh_Alarm[11].Healthy, AlarmOut => "1092_HMI_OP_FLAGS".LS425_442_LevelSwitch_HighHigh_Alarm[11].UnhealthyAlarm)
   END_RUNG
   // the same network as SCL:
   "1602_DIGITAL_HEALTH"(InputSignal := "20_TANKS_IP_DATA".RIO_05.FIRST_TANK.BWT_LEVEL_HIHI,
                         InputTripLevel := #InputTripLevel,
                         SensorHealthOut => "1092_HMI_OP_FLAGS".LS425_442_LevelSwitch_HighHigh_Alarm[10].Healthy,
                         AlarmOut => "1092_HMI_OP_FLAGS".LS425_442_LevelSwitch_HighHigh_Alarm[10].UnhealthyAlarm);
   "1602_DIGITAL_HEALTH"(InputSignal := "20_TANKS_IP_DATA".RIO_05.SECOND_TANK.BWT_LEVEL_HIHI,
                         InputTripLevel := #InputTripLevel,
                         SensorHealthOut => "1092_HMI_OP_FLAGS".LS425_442_LevelSwitch_HighHigh_Alarm[11].Healthy,
                         AlarmOut => "1092_HMI_OP_FLAGS".LS425_442_LevelSwitch_HighHigh_Alarm[11].UnhealthyAlarm);
END_REGION

REGION Network 6: LS425, LS442 Alarms (RIO 06: 6P, 6S)
   RUNG wire#powerrail
      "1602_DIGITAL_HEALTH"(InputSignal := "20_TANKS_IP_DATA".RIO_06.FIRST_TANK.BWT_LEVEL_HIHI, InputTripLevel := #InputTripLevel, SensorHealthOut => "1092_HMI_OP_FLAGS".LS425_442_LevelSwitch_HighHigh_Alarm[12].Healthy, AlarmOut => "1092_HMI_OP_FLAGS".LS425_442_LevelSwitch_HighHigh_Alarm[12].UnhealthyAlarm)
   END_RUNG
   RUNG wire#powerrail
      "1602_DIGITAL_HEALTH"(InputSignal := "20_TANKS_IP_DATA".RIO_06.SECOND_TANK.BWT_LEVEL_HIHI, InputTripLevel := #InputTripLevel, SensorHealthOut => "1092_HMI_OP_FLAGS".LS425_442_LevelSwitch_HighHigh_Alarm[13].Healthy, AlarmOut => "1092_HMI_OP_FLAGS".LS425_442_LevelSwitch_HighHigh_Alarm[13].UnhealthyAlarm)
   END_RUNG
   // the same network as SCL:
   "1602_DIGITAL_HEALTH"(InputSignal := "20_TANKS_IP_DATA".RIO_06.FIRST_TANK.BWT_LEVEL_HIHI,
                         InputTripLevel := #InputTripLevel,
                         SensorHealthOut => "1092_HMI_OP_FLAGS".LS425_442_LevelSwitch_HighHigh_Alarm[12].Healthy,
                         AlarmOut => "1092_HMI_OP_FLAGS".LS425_442_LevelSwitch_HighHigh_Alarm[12].UnhealthyAlarm);
   "1602_DIGITAL_HEALTH"(InputSignal := "20_TANKS_IP_DATA".RIO_06.SECOND_TANK.BWT_LEVEL_HIHI,
                         InputTripLevel := #InputTripLevel,
                         SensorHealthOut => "1092_HMI_OP_FLAGS".LS425_442_LevelSwitch_HighHigh_Alarm[13].Healthy,
                         AlarmOut => "1092_HMI_OP_FLAGS".LS425_442_LevelSwitch_HighHigh_Alarm[13].UnhealthyAlarm);
END_REGION

